        [84].runs[11] := 9, [84].runs[12] := 9, [84].runs[13] := 9, [84].runs[14] := 9, [84].runs[15] := 10, [84].runs[16] := 9, [84].runs[17] := 10, [84].runs[18] := 9, [84].runs[19] := 10, [84].runs[20] := 9, [84].runs[21] := 8, [84].runs[22] := 5, [84].time_avg[0] := 173, [84].time_avg[2] := 6434, [84].time_avg[3] := 9546, [84].time_avg[4] := 19840, [84].time_avg[5] := 19601, [84].time_avg[10] := 183, [84].time_avg[11] := 176, [84].time_avg[12] := 189, [84].time_avg[13] := 198, [84].time_avg[14] := 193, [84].time_avg[15] := 154, [84].time_avg[16] := 205, [84].time_avg[17] := 165, [84].time_avg[18] := 168, [84].time_avg[19] := 167, [84].time_avg[20] := 143, [84].time_avg[21] := 164, [84].time_avg[22] := 139, [85].date[0] := 19, [85].date[1] := 8, [85].date[2] := 23, [85].runs[0] := 108, [85].runs[7] := 1, [85].runs[9] := 4, [85].runs[10] := 3, [85].runs[11] := 10, [85].runs[12] := 9, [85].runs[13] := 8, [85].runs[14] := 9, [85].runs[15] := 10, [85].runs[16] := 9, [85].runs[17] := 9, [85].runs[18] := 8, [85].runs[19] := 9, [85].runs[20] := 9, [85].runs[21] := 8, [85].runs[22] := 2, [85].time_avg[0] := 204, [85].time_avg[2] := 6887, [85].time_avg[3] := 14477, [85].time_avg[4] := 20521, [85].time_avg[5] := 36240, [85].time_avg[10] := 221, [85].time_avg[11] := 190, [85].time_avg[12] := 186, [85].time_avg[13] := 191, [85].time_avg[14] := 226, [85].time_avg[15] := 161,
        [85].time_avg[16] := 185, [85].time_avg[17] := 211, [85].time_avg[18] := 232, [85].time_avg[19] := 218, [85].time_avg[20] := 196, [85].time_avg[21] := 251, [85].time_avg[22] := 235, [86].date[0] := 19, [86].date[1] := 8, [86].date[2] := 22, [86].runs[0] := 108, [86].runs[9] := 4, [86].runs[10] := 5, [86].runs[11] := 10, [86].runs[12] := 9, [86].runs[13] := 11, [86].runs[14] := 9, [86].runs[15] := 10, [86].runs[16] := 9, [86].runs[17] := 10, [86].runs[18] := 8, [86].runs[19] := 10, [86].runs[20] := 9, [86].runs[21] := 3, [86].time_avg[0] := 162, [86].time_avg[2] := 5022, [86].time_avg[3] := 11042, [86].time_avg[4] := 16840, [86].time_avg[5] := 22478, [86].time_avg[10] := 152, [86].time_avg[11] := 173, [86].time_avg[12] := 166, [86].time_avg[13] := 153, [86].time_avg[14] := 137, [86].time_avg[15] := 192, [86].time_avg[16] := 160, [86].time_avg[17] := 147, [86].time_avg[18] := 177, [86].time_avg[19] := 145, [86].time_avg[20] := 166, [86].time_avg[21] := 190, [87].date[0] := 19, [87].date[1] := 8, [87].date[2] := 21, [87].runs[0] := 110, [87].runs[9] := 5, [87].runs[10] := 5, [87].runs[11] := 9, [87].runs[12] := 8, [87].runs[13] := 10, [87].runs[14] := 10, [87].runs[15] := 10, [87].runs[16] := 10, [87].runs[17] := 9, [87].runs[18] := 10, [87].runs[19] := 8, [87].runs[20] := 9, [87].runs[21] := 6, [87].time_avg[0] := 174, [87].time_avg[2] := 5028,
        [87].time_avg[3] := 12622, [87].time_avg[4] := 18641, [87].time_avg[5] := 20757, [87].time_avg[9] := 267, [87].time_avg[10] := 158, [87].time_avg[11] := 186, [87].time_avg[12] := 162, [87].time_avg[13] := 179, [87].time_avg[14] := 156, [87].time_avg[15] := 147, [87].time_avg[16] := 154, [87].time_avg[17] := 158, [87].time_avg[18] := 185, [87].time_avg[19] := 180, [87].time_avg[20] := 236, [87].time_avg[21] := 167, [88].date[0] := 19, [88].date[1] := 8, [88].date[2] := 19, [88].runs[0] := 172, [88].runs[7] := 1, [88].runs[9] := 1, [88].runs[10] := 7, [88].runs[11] := 9, [88].runs[12] := 10, [88].runs[13] := 10, [88].runs[14] := 10, [88].runs[15] := 10, [88].runs[16] := 9, [88].runs[17] := 9, [88].runs[18] := 10, [88].runs[19] := 11, [88].runs[20] := 10, [88].runs[21] := 8, [88].time_avg[0] := 159, [88].time_avg[2] := 5010, [88].time_avg[3] := 9465, [88].time_avg[4] := 20080, [88].time_avg[5] := 17563, [88].time_avg[10] := 264, [88].time_avg[11] := 192, [88].time_avg[12] := 158, [88].time_avg[13] := 167, [88].time_avg[14] := 165, [88].time_avg[15] := 148, [88].time_avg[16] := 206, [88].time_avg[17] := 174, [88].time_avg[18] := 142, [88].time_avg[19] := 133, [88].time_avg[20] := 165, [88].time_avg[21] := 129, [89].date[0] := 19, [89].date[1] := 8, [89].date[2] := 18, [89].runs[0] := 116, [89].runs[7] := 1, [89].runs[10] := 8, [89].runs[11] := 10, [89].runs[12] := 10, [89].runs[13] := 9,
        [89].runs[14] := 10, [89].runs[15] := 11, [89].runs[16] := 4, [89].runs[17] := 9, [89].runs[18] := 10, [89].runs[19] := 10, [89].runs[20] := 9, [89].runs[21] := 11, [89].runs[22] := 4, [89].time_avg[0] := 160, [89].time_avg[2] := 4655, [89].time_avg[3] := 12877, [89].time_avg[4] := 21363, [89].time_avg[5] := 26439, [89].time_avg[10] := 166, [89].time_avg[11] := 166, [89].time_avg[12] := 161, [89].time_avg[13] := 187, [89].time_avg[14] := 165, [89].time_avg[15] := 133, [89].time_avg[16] := 160, [89].time_avg[17] := 161, [89].time_avg[18] := 173, [89].time_avg[19] := 149, [89].time_avg[20] := 175, [89].time_avg[21] := 139, [89].time_avg[22] := 162, [90].date[0] := 19, [90].date[1] := 8, [90].date[2] := 17, [90].runs[0] := 129, [90].runs[7] := 1, [90].runs[9] := 4, [90].runs[10] := 4, [90].runs[11] := 10, [90].runs[12] := 9, [90].runs[13] := 10, [90].runs[14] := 10, [90].runs[15] := 9, [90].runs[16] := 10, [90].runs[17] := 10, [90].runs[18] := 7, [90].runs[19] := 9, [90].runs[20] := 8, [90].runs[21] := 9, [90].runs[22] := 10, [90].runs[23] := 8, [90].time_avg[0] := 182, [90].time_avg[2] := 4196, [90].time_avg[3] := 11369, [90].time_avg[4] := 22122, [90].time_avg[5] := 21841, [90].time_avg[10] := 197, [90].time_avg[11] := 174, [90].time_avg[12] := 191, [90].time_avg[13] := 174, [90].time_avg[14] := 150, [90].time_avg[15] := 171, [90].time_avg[16] := 159, [90].time_avg[17] := 162,
        [90].time_avg[18] := 179, [90].time_avg[19] := 213, [90].time_avg[20] := 216, [90].time_avg[21] := 192, [90].time_avg[22] := 182, [90].time_avg[23] := 211, [91].date[0] := 19, [91].date[1] := 8, [91].date[2] := 16, [91].runs[0] := 110, [91].runs[7] := 1, [91].runs[9] := 4, [91].runs[10] := 6, [91].runs[11] := 10, [91].runs[12] := 8, [91].runs[13] := 9, [91].runs[14] := 3, [91].runs[15] := 10, [91].runs[16] := 10, [91].runs[17] := 10, [91].runs[18] := 9, [91].runs[19] := 9, [91].runs[20] := 9, [91].runs[21] := 10, [91].runs[22] := 2, [91].time_avg[0] := 167, [91].time_avg[2] := 5926, [91].time_avg[3] := 9632, [91].time_avg[4] := 23480, [91].time_avg[5] := 18838, [91].time_avg[10] := 161, [91].time_avg[11] := 149, [91].time_avg[12] := 156, [91].time_avg[13] := 170, [91].time_avg[15] := 151, [91].time_avg[16] := 156, [91].time_avg[17] := 158, [91].time_avg[18] := 203, [91].time_avg[19] := 192, [91].time_avg[20] := 185, [91].time_avg[21] := 150, [91].time_avg[22] := 195, [92].date[0] := 19, [92].date[1] := 8, [92].date[2] := 15, [92].runs[0] := 113, [92].runs[7] := 1, [92].runs[9] := 4, [92].runs[10] := 5, [92].runs[11] := 9, [92].runs[12] := 9, [92].runs[13] := 9, [92].runs[14] := 9, [92].runs[15] := 10, [92].runs[16] := 10, [92].runs[17] := 9, [92].runs[18] := 10, [92].runs[19] := 9, [92].runs[20] := 10, [92].runs[21] := 9,
        [92].time_avg[0] := 174, [92].time_avg[2] := 4980, [92].time_avg[3] := 11102, [92].time_avg[4] := 19122, [92].time_avg[5] := 22677, [92].time_avg[10] := 180, [92].time_avg[11] := 184, [92].time_avg[12] := 201, [92].time_avg[13] := 188, [92].time_avg[14] := 179, [92].time_avg[15] := 164, [92].time_avg[16] := 165, [92].time_avg[17] := 189, [92].time_avg[18] := 169, [92].time_avg[19] := 168, [92].time_avg[20] := 159, [92].time_avg[21] := 153, [93].date[0] := 19, [93].date[1] := 8, [93].date[2] := 14, [93].runs[0] := 110, [93].runs[7] := 1, [93].runs[9] := 4, [93].runs[10] := 5, [93].runs[11] := 9, [93].runs[12] := 10, [93].runs[13] := 10, [93].runs[14] := 10, [93].runs[15] := 10, [93].runs[16] := 10, [93].runs[17] := 8, [93].runs[18] := 10, [93].runs[19] := 10, [93].runs[20] := 8, [93].runs[21] := 5, [93].time_avg[0] := 170, [93].time_avg[2] := 3396, [93].time_avg[3] := 11574, [93].time_avg[4] := 19402, [93].time_avg[5] := 24403, [93].time_avg[10] := 164, [93].time_avg[11] := 183, [93].time_avg[12] := 161, [93].time_avg[13] := 163, [93].time_avg[14] := 151, [93].time_avg[15] := 150, [93].time_avg[16] := 168, [93].time_avg[17] := 227, [93].time_avg[18] := 179, [93].time_avg[19] := 161, [93].time_avg[20] := 173, [93].time_avg[21] := 178, [94].date[0] := 19, [94].date[1] := 8, [94].date[2] := 13, [94].runs[0] := 99, [94].runs[7] := 1, [94].runs[9] := 4, [94].runs[10] := 4, [94].runs[11] := 11,
        [94].runs[12] := 8, [94].runs[13] := 5, [94].runs[14] := 9, [94].runs[15] := 8, [94].runs[16] := 10, [94].runs[17] := 9, [94].runs[18] := 8, [94].runs[19] := 9, [94].runs[20] := 8, [94].runs[21] := 5, [94].time_avg[0] := 185, [94].time_avg[2] := 4905, [94].time_avg[3] := 9992, [94].time_avg[4] := 19077, [94].time_avg[5] := 20762, [94].time_avg[10] := 183, [94].time_avg[11] := 135, [94].time_avg[12] := 171, [94].time_avg[13] := 195, [94].time_avg[14] := 209, [94].time_avg[15] := 185, [94].time_avg[16] := 185, [94].time_avg[17] := 186, [94].time_avg[18] := 200, [94].time_avg[19] := 175, [94].time_avg[20] := 224, [94].time_avg[21] := 204, [95].date[0] := 19, [95].date[1] := 8, [95].date[2] := 12, [95].runs[0] := 118, [95].runs[8] := 1, [95].runs[9] := 6, [95].runs[10] := 5, [95].runs[11] := 10, [95].runs[12] := 11, [95].runs[13] := 10, [95].runs[14] := 8, [95].runs[15] := 10, [95].runs[16] := 10, [95].runs[17] := 10, [95].runs[18] := 10, [95].runs[19] := 8, [95].runs[20] := 9, [95].runs[21] := 10, [95].time_avg[0] := 156, [95].time_avg[2] := 6366, [95].time_avg[3] := 11660, [95].time_avg[4] := 23243, [95].time_avg[5] := 28239, [95].time_avg[10] := 194, [95].time_avg[11] := 153, [95].time_avg[12] := 133, [95].time_avg[13] := 156, [95].time_avg[14] := 137, [95].time_avg[15] := 150, [95].time_avg[16] := 151, [95].time_avg[17] := 145, [95].time_avg[18] := 164, [95].time_avg[19] := 182,
        [95].time_avg[20] := 195, [95].time_avg[21] := 148, [96].date[0] := 19, [96].date[1] := 8, [96].date[2] := 11, [96].runs[0] := 123, [96].runs[7] := 1, [96].runs[9] := 4, [96].runs[10] := 8, [96].runs[11] := 10, [96].runs[12] := 11, [96].runs[13] := 10, [96].runs[14] := 7, [96].runs[15] := 11, [96].runs[16] := 9, [96].runs[17] := 10, [96].runs[18] := 9, [96].runs[19] := 11, [96].runs[20] := 8, [96].runs[21] := 9, [96].runs[22] := 5, [96].time_avg[0] := 157, [96].time_avg[2] := 4752, [96].time_avg[3] := 9692, [96].time_avg[4] := 19361, [96].time_avg[5] := 22281, [96].time_avg[10] := 173, [96].time_avg[11] := 141, [96].time_avg[12] := 142, [96].time_avg[13] := 141, [96].time_avg[14] := 179, [96].time_avg[15] := 138, [96].time_avg[16] := 183, [96].time_avg[17] := 147, [96].time_avg[18] := 191, [96].time_avg[19] := 146, [96].time_avg[20] := 167, [96].time_avg[21] := 162, [96].time_avg[22] := 167, [97].date[0] := 19, [97].date[1] := 8, [97].date[2] := 10, [97].runs[0] := 120, [97].runs[7] := 1, [97].runs[9] := 5, [97].runs[10] := 4, [97].runs[11] := 6, [97].runs[12] := 8, [97].runs[13] := 11, [97].runs[14] := 8, [97].runs[15] := 11, [97].runs[16] := 9, [97].runs[17] := 10, [97].runs[18] := 11, [97].runs[19] := 10, [97].runs[20] := 11, [97].runs[21] := 10, [97].runs[22] := 5, [97].time_avg[0] := 142, [97].time_avg[2] := 4697,
        [97].time_avg[3] := 8479, [97].time_avg[4] := 21362, [97].time_avg[5] := 36560, [97].time_avg[10] := 200, [97].time_avg[11] := 178, [97].time_avg[12] := 152, [97].time_avg[13] := 141, [97].time_avg[14] := 131, [97].time_avg[15] := 153, [97].time_avg[16] := 133, [97].time_avg[17] := 145, [97].time_avg[18] := 140, [97].time_avg[19] := 135, [97].time_avg[20] := 138, [97].time_avg[21] := 126, [97].time_avg[22] := 121, [98].date[0] := 19, [98].date[1] := 8, [98].date[2] := 9, [98].runs[0] := 119, [98].runs[7] := 1, [98].runs[9] := 5, [98].runs[10] := 5, [98].runs[11] := 8, [98].runs[12] := 9, [98].runs[13] := 8, [98].runs[14] := 11, [98].runs[15] := 11, [98].runs[16] := 8, [98].runs[17] := 10, [98].runs[18] := 9, [98].runs[19] := 11, [98].runs[20] := 9, [98].runs[21] := 10, [98].runs[22] := 4, [98].time_avg[0] := 151, [98].time_avg[2] := 4804, [98].time_avg[3] := 10881, [98].time_avg[4] := 800, [98].time_avg[5] := 21920, [98].time_avg[9] := 35, [98].time_avg[10] := 126, [98].time_avg[11] := 166, [98].time_avg[12] := 159, [98].time_avg[13] := 165, [98].time_avg[14] := 138, [98].time_avg[15] := 126, [98].time_avg[16] := 148, [98].time_avg[17] := 148, [98].time_avg[18] := 187, [98].time_avg[19] := 138, [98].time_avg[20] := 165, [98].time_avg[21] := 145, [98].time_avg[22] := 168, [99].date[0] := 19, [99].date[1] := 8, [99].date[2] := 8, [99].runs[0] := 93, [99].runs[7] := 1, [99].runs[9] := 4,
        [99].runs[10] := 4, [99].runs[11] := 9, [99].runs[12] := 9, [99].runs[13] := 9, [99].runs[14] := 8, [99].runs[15] := 9, [99].runs[16] := 9, [99].runs[17] := 2, [99].runs[18] := 5, [99].runs[19] := 8, [99].runs[20] := 9, [99].runs[21] := 7, [99].time_avg[0] := 156, [99].time_avg[2] := 5998, [99].time_avg[3] := 7111, [99].time_avg[4] := 17880, [99].time_avg[5] := 21321, [99].time_avg[10] := 153, [99].time_avg[11] := 154, [99].time_avg[12] := 146, [99].time_avg[13] := 139, [99].time_avg[14] := 173, [99].time_avg[15] := 152, [99].time_avg[16] := 160, [99].time_avg[17] := 133, [99].time_avg[18] := 182, [99].time_avg[19] := 147, [99].time_avg[20] := 148, [99].time_avg[21] := 188);
        [0].time_avg[2]   // Daily Avg Platform Cycle Waiting After Cycle
        [0].time_avg[3]   // Daily Avg Platform Cycle Before Start Cycle
        [0].time_avg[4]   // Overall Time End of Cycle Plat
        [0].time_avg[5]   // Overall Time Before Cycle Plat
   JM_Statistics_Storage : Run_Count_Hist_JM[100] := ([1].date[0] := 25, [1].date[1] := 11, [1].date[2] := 28, [1].runs[0] := 65, [1].runs[8] := 2, [1].runs[9] := 1, [1].runs[15] := 3, [1].runs[16] := 7, [1].runs[17] := 8, [1].runs[18] := 8, [1].runs[19] := 8, [1].runs[20] := 8, [1].runs[21] := 7, [1].runs[22] := 8, [1].runs[23] := 5, [1].time_avg[0] := 204, [1].time_avg[2] := 3400, [1].time_avg[4] := 19639, [1].time_avg[5] := 22361, [1].time_avg[8] := 50, [1].time_avg[15] := 203, [1].time_avg[16] := 254, [1].time_avg[17] := 210, [1].time_avg[18] := 202, [1].time_avg[19] := 195, [1].time_avg[20] := 206, [1].time_avg[21] := 190, [1].time_avg[22] := 211, [1].time_avg[23] := 177, [2].date[0] := 25, [2].date[1] := 11, [2].date[2] := 27, [2].runs[0] := 63, [2].runs[14] := 6, [2].runs[15] := 4, [2].runs[16] := 7, [2].runs[17] := 7, [2].runs[18] := 8, [2].runs[19] := 8, [2].runs[20] := 7, [2].runs[21] := 5, [2].runs[22] := 8, [2].runs[23] := 3, [2].time_avg[0] := 234, [2].time_avg[4] := 21760, [2].time_avg[5] := 22361, [2].time_avg[14] := 167, [2].time_avg[15] := 316, [2].time_avg[16] := 272, [2].time_avg[17] := 206, [2].time_avg[18] := 208, [2].time_avg[19] := 242, [2].time_avg[20] := 266, [2].time_avg[21] := 233, [2].time_avg[22] := 223, [2].time_avg[23] := 245, [3].date[0] := 25, [3].date[1] := 11, [3].date[2] := 26, [3].runs[0] := 57,
        [3].runs[12] := 4, [3].runs[13] := 1, [3].runs[15] := 2, [3].runs[16] := 6, [3].runs[17] := 7, [3].runs[18] := 7, [3].runs[19] := 7, [3].runs[20] := 7, [3].runs[21] := 7, [3].runs[22] := 6, [3].runs[23] := 3, [3].time_avg[0] := 274, [3].time_avg[2] := 6041, [3].time_avg[4] := 21760, [3].time_avg[5] := 22361, [3].time_avg[12] := 396, [3].time_avg[13] := 320, [3].time_avg[15] := 271, [3].time_avg[16] := 271, [3].time_avg[17] := 292, [3].time_avg[18] := 243, [3].time_avg[19] := 255, [3].time_avg[20] := 243, [3].time_avg[21] := 289, [3].time_avg[22] := 278, [3].time_avg[23] := 283, [4].date[0] := 25, [4].date[1] := 11, [4].date[2] := 25, [4].runs[0] := 53, [4].runs[7] := 1, [4].runs[15] := 1, [4].runs[16] := 5, [4].runs[17] := 8, [4].runs[18] := 6, [4].runs[19] := 8, [4].runs[20] := 7, [4].runs[21] := 7, [4].runs[22] := 7, [4].runs[23] := 3, [4].time_avg[0] := 260, [4].time_avg[4] := 53080, [4].time_avg[5] := 22361, [4].time_avg[16] := 223, [4].time_avg[17] := 286, [4].time_avg[18] := 280, [4].time_avg[19] := 258, [4].time_avg[20] := 261, [4].time_avg[21] := 234, [4].time_avg[22] := 267, [4].time_avg[23] := 254, [5].date[0] := 25, [5].date[1] := 11, [5].date[2] := 24, [5].runs[0] := 67, [5].runs[7] := 4, [5].runs[8] := 3, [5].runs[10] := 2, [5].runs[11] := 4, [5].runs[13] := 1,
        [5].runs[14] := 1, [5].runs[15] := 4, [5].runs[16] := 7, [5].runs[17] := 7, [5].runs[18] := 7, [5].runs[19] := 7, [5].runs[20] := 4, [5].runs[21] := 7, [5].runs[22] := 6, [5].runs[23] := 3, [5].time_avg[0] := 254, [5].time_avg[2] := 76642, [5].time_avg[4] := 53080, [5].time_avg[5] := 22361, [5].time_avg[7] := 75, [5].time_avg[8] := 246, [5].time_avg[11] := 171, [5].time_avg[14] := 83, [5].time_avg[15] := 147, [5].time_avg[16] := 272, [5].time_avg[17] := 276, [5].time_avg[18] := 244, [5].time_avg[19] := 256, [5].time_avg[20] := 266, [5].time_avg[21] := 291, [5].time_avg[22] := 291, [5].time_avg[23] := 290, [6].date[0] := 25, [6].date[1] := 11, [6].date[2] := 23, [6].runs[0] := 54, [6].runs[10] := 2, [6].runs[11] := 4, [6].runs[15] := 1, [6].runs[16] := 8, [6].runs[17] := 7, [6].runs[18] := 6, [6].runs[19] := 5, [6].runs[20] := 8, [6].runs[21] := 6, [6].runs[22] := 5, [6].runs[23] := 2, [6].time_avg[0] := 268, [6].time_avg[4] := 23760, [6].time_avg[5] := 22361, [6].time_avg[11] := 332, [6].time_avg[16] := 211, [6].time_avg[17] := 253, [6].time_avg[18] := 262, [6].time_avg[19] := 274, [6].time_avg[20] := 241, [6].time_avg[21] := 295, [6].time_avg[22] := 310, [6].time_avg[23] := 371, [7].date[0] := 25, [7].date[1] := 11, [7].date[2] := 22, [7].runs[0] := 49, [7].runs[12] := 7, [7].runs[14] := 1,
        [7].runs[15] := 4, [7].runs[16] := 7, [7].runs[17] := 7, [7].runs[18] := 7, [7].runs[19] := 1, [7].runs[20] := 6, [7].runs[21] := 2, [7].runs[22] := 6, [7].runs[23] := 1, [7].time_avg[0] := 278, [7].time_avg[4] := 23760, [7].time_avg[5] := 22361, [7].time_avg[12] := 180, [7].time_avg[15] := 308, [7].time_avg[16] := 282, [7].time_avg[17] := 261, [7].time_avg[18] := 280, [7].time_avg[19] := 295, [7].time_avg[20] := 361, [7].time_avg[22] := 287, [8].date[0] := 25, [8].date[1] := 11, [8].date[2] := 20, [8].runs[0] := 58, [8].runs[10] := 2, [8].runs[11] := 3, [8].runs[13] := 5, [8].runs[14] := 4, [8].runs[15] := 3, [8].runs[16] := 5, [8].runs[17] := 4, [8].runs[18] := 3, [8].runs[19] := 6, [8].runs[20] := 5, [8].runs[21] := 7, [8].runs[22] := 7, [8].runs[23] := 4, [8].time_avg[0] := 205, [8].time_avg[2] := 15381, [8].time_avg[4] := 23760, [8].time_avg[5] := 22361, [8].time_avg[10] := 76, [8].time_avg[11] := 152, [8].time_avg[13] := 198, [8].time_avg[14] := 60, [8].time_avg[15] := 73, [8].time_avg[16] := 76, [8].time_avg[17] := 183, [8].time_avg[18] := 376, [8].time_avg[19] := 286, [8].time_avg[20] := 250, [8].time_avg[21] := 218, [8].time_avg[22] := 239, [8].time_avg[23] := 211, [9].date[0] := 25, [9].date[1] := 11, [9].date[2] := 19, [9].runs[0] := 7, [9].runs[12] := 2, [9].runs[13] := 4,
        [9].runs[17] := 1, [9].runs[18] := 1, [9].time_avg[0] := 217, [9].time_avg[2] := 78801, [9].time_avg[4] := 48480, [9].time_avg[5] := 22361, [9].time_avg[13] := 217, [10].date[0] := 25, [10].date[1] := 11, [10].date[2] := 16, [10].runs[0] := 7, [10].runs[10] := 2, [10].runs[13] := 7, [10].time_avg[0] := 93, [10].time_avg[4] := 27759, [10].time_avg[5] := 22361, [10].time_avg[13] := 93, [11].date[0] := 25, [11].date[1] := 11, [11].date[2] := 14, [11].runs[0] := 2, [11].runs[15] := 1, [11].runs[16] := 1, [11].time_avg[2] := 32760, [11].time_avg[4] := 27759, [11].time_avg[5] := 22361, [12].date[0] := 25, [12].date[1] := 11, [12].date[2] := 13, [12].runs[0] := 14, [12].runs[10] := 2, [12].runs[11] := 1, [12].runs[12] := 1, [12].runs[14] := 2, [12].runs[15] := 5, [12].runs[16] := 4, [12].runs[17] := 5, [12].time_avg[0] := 141, [12].time_avg[4] := 36240, [12].time_avg[5] := 22361, [12].time_avg[10] := 210, [12].time_avg[14] := 205, [12].time_avg[15] := 160, [12].time_avg[16] := 100, [12].time_avg[17] := 100, [13].date[0] := 25, [13].date[1] := 11, [13].date[2] := 11, [13].runs[0] := 2, [13].runs[18] := 2, [13].time_avg[0] := 88, [13].time_avg[4] := 36240, [13].time_avg[5] := 22361, [13].time_avg[18] := 88, [14].date[0] := 25, [14].date[1] := 11, [14].date[2] := 7, [14].runs[0] := 5, [14].runs[15] := 3, [14].runs[16] := 2,
        [14].time_avg[0] := 229, [14].time_avg[4] := 36240, [14].time_avg[5] := 22361, [14].time_avg[15] := 300, [14].time_avg[16] := 87, [15].date[0] := 25, [15].date[1] := 11, [15].date[2] := 6, [15].runs[0] := 13, [15].runs[15] := 1, [15].runs[16] := 3, [15].runs[17] := 8, [15].runs[18] := 1, [15].runs[19] := 4, [15].time_avg[0] := 54, [15].time_avg[4] := 36240, [15].time_avg[5] := 22361, [15].time_avg[17] := 46, [15].time_avg[19] := 66, [16].date[0] := 25, [16].date[1] := 10, [16].date[2] := 27, [16].runs[0] := 13, [16].runs[12] := 1, [16].runs[13] := 4, [16].runs[14] := 1, [16].time_avg[0] := 126, [16].time_avg[4] := 36240, [16].time_avg[5] := 22361, [16].time_avg[13] := 65, [17].date[0] := 25, [17].date[1] := 10, [17].date[2] := 26, [17].runs[0] := 58, [17].runs[10] := 1, [17].runs[11] := 2, [17].runs[12] := 3, [17].runs[13] := 8, [17].runs[14] := 8, [17].runs[15] := 6, [17].runs[16] := 7, [17].runs[17] := 7, [17].runs[18] := 6, [17].runs[19] := 7, [17].runs[20] := 3, [17].time_avg[0] := 252, [17].time_avg[2] := 40720, [17].time_avg[4] := 36240, [17].time_avg[5] := 22361, [17].time_avg[11] := 476, [17].time_avg[12] := 190, [17].time_avg[13] := 206, [17].time_avg[14] := 216, [17].time_avg[15] := 310, [17].time_avg[16] := 261, [17].time_avg[17] := 248, [17].time_avg[18] := 232, [17].time_avg[19] := 304, [17].time_avg[20] := 214, [18].date[0] := 25,
        [18].date[1] := 10, [18].date[2] := 25, [18].runs[0] := 47, [18].runs[12] := 5, [18].runs[13] := 9, [18].runs[14] := 5, [18].runs[16] := 2, [18].runs[17] := 8, [18].runs[18] := 7, [18].runs[19] := 7, [18].runs[20] := 4, [18].time_avg[0] := 227, [18].time_avg[4] := 26040, [18].time_avg[5] := 22361, [18].time_avg[12] := 203, [18].time_avg[13] := 166, [18].time_avg[14] := 231, [18].time_avg[16] := 370, [18].time_avg[17] := 239, [18].time_avg[18] := 252, [18].time_avg[19] := 244, [18].time_avg[20] := 235, [19].date[0] := 25, [19].date[1] := 10, [19].date[2] := 23, [19].runs[0] := 48, [19].runs[9] := 2, [19].runs[10] := 3, [19].runs[12] := 3, [19].runs[13] := 7, [19].runs[14] := 7, [19].runs[15] := 5, [19].runs[16] := 8, [19].runs[17] := 5, [19].runs[19] := 5, [19].runs[20] := 3, [19].time_avg[0] := 257, [19].time_avg[2] := 18201, [19].time_avg[4] := 26040, [19].time_avg[5] := 22361, [19].time_avg[9] := 102, [19].time_avg[10] := 259, [19].time_avg[12] := 493, [19].time_avg[13] := 241, [19].time_avg[14] := 231, [19].time_avg[15] := 264, [19].time_avg[16] := 252, [19].time_avg[17] := 280, [19].time_avg[19] := 300, [19].time_avg[20] := 235, [20].date[0] := 25, [20].date[1] := 10, [20].date[2] := 22, [20].runs[0] := 62, [20].runs[10] := 4, [20].runs[12] := 2, [20].runs[13] := 9, [20].runs[14] := 7, [20].runs[15] := 7, [20].runs[16] := 7,
        [20].runs[17] := 7, [20].runs[18] := 8, [20].runs[19] := 8, [20].runs[20] := 3, [20].time_avg[0] := 226, [20].time_avg[4] := 26079, [20].time_avg[5] := 22361, [20].time_avg[10] := 123, [20].time_avg[13] := 199, [20].time_avg[14] := 230, [20].time_avg[15] := 230, [20].time_avg[16] := 312, [20].time_avg[17] := 253, [20].time_avg[18] := 219, [20].time_avg[19] := 200, [20].time_avg[20] := 206, [21].date[0] := 25, [21].date[1] := 10, [21].date[2] := 21, [21].runs[0] := 58, [21].runs[11] := 3, [21].runs[12] := 1, [21].runs[13] := 8, [21].runs[14] := 7, [21].runs[15] := 4, [21].runs[16] := 8, [21].runs[17] := 8, [21].runs[18] := 7, [21].runs[19] := 8, [21].runs[20] := 4, [21].time_avg[0] := 233, [21].time_avg[2] := 42160, [21].time_avg[4] := 26079, [21].time_avg[5] := 22361, [21].time_avg[11] := 186, [21].time_avg[13] := 222, [21].time_avg[14] := 240, [21].time_avg[15] := 294, [21].time_avg[16] := 256, [21].time_avg[17] := 202, [21].time_avg[18] := 246, [21].time_avg[19] := 216, [21].time_avg[20] := 208, [22].date[0] := 25, [22].date[1] := 10, [22].date[2] := 20, [22].runs[0] := 47, [22].runs[10] := 2, [22].runs[11] := 6, [22].runs[12] := 1, [22].runs[13] := 7, [22].runs[14] := 7, [22].runs[15] := 7, [22].runs[16] := 4, [22].runs[17] := 1, [22].runs[18] := 2, [22].runs[19] := 7, [22].runs[20] := 3, [22].time_avg[0] := 249, [22].time_avg[2] := 52640,
        [22].time_avg[4] := 40960, [22].time_avg[5] := 22361, [22].time_avg[11] := 232, [22].time_avg[13] := 215, [22].time_avg[14] := 258, [22].time_avg[15] := 237, [22].time_avg[16] := 210, [22].time_avg[18] := 331, [22].time_avg[19] := 294, [22].time_avg[20] := 241, [23].date[0] := 25, [23].date[1] := 10, [23].date[2] := 19, [23].runs[0] := 61, [23].runs[9] := 2, [23].runs[10] := 2, [23].runs[11] := 8, [23].runs[12] := 4, [23].runs[13] := 6, [23].runs[14] := 1, [23].runs[15] := 8, [23].runs[16] := 7, [23].runs[17] := 7, [23].runs[18] := 7, [23].runs[19] := 7, [23].runs[20] := 2, [23].time_avg[0] := 237, [23].time_avg[2] := 59762, [23].time_avg[4] := 52320, [23].time_avg[5] := 22361, [23].time_avg[9] := 89, [23].time_avg[11] := 203, [23].time_avg[12] := 193, [23].time_avg[13] := 194, [23].time_avg[15] := 243, [23].time_avg[16] := 238, [23].time_avg[17] := 251, [23].time_avg[18] := 268, [23].time_avg[19] := 280, [23].time_avg[20] := 287, [24].date[0] := 25, [24].date[1] := 10, [24].date[2] := 18, [24].runs[0] := 51, [24].runs[9] := 2, [24].runs[10] := 5, [24].runs[11] := 8, [24].runs[12] := 2, [24].runs[13] := 5, [24].runs[14] := 6, [24].runs[15] := 7, [24].runs[16] := 5, [24].runs[17] := 7, [24].runs[18] := 4, [24].time_avg[0] := 246, [24].time_avg[4] := 52360, [24].time_avg[5] := 22361, [24].time_avg[10] := 182, [24].time_avg[11] := 228, [24].time_avg[12] := 212,
        [24].time_avg[13] := 231, [24].time_avg[14] := 324, [24].time_avg[15] := 255, [24].time_avg[16] := 238, [24].time_avg[17] := 263, [24].time_avg[18] := 255, [25].date[0] := 25, [25].date[1] := 10, [25].date[2] := 15, [25].runs[0] := 89, [25].runs[10] := 4, [25].runs[11] := 4, [25].runs[12] := 7, [25].runs[13] := 6, [25].runs[14] := 8, [25].runs[15] := 6, [25].runs[16] := 7, [25].runs[17] := 6, [25].time_avg[0] := 251, [25].time_avg[2] := 50482, [25].time_avg[4] := 52360, [25].time_avg[5] := 22361, [25].time_avg[10] := 61, [25].time_avg[11] := 214, [25].time_avg[12] := 261, [25].time_avg[13] := 348, [25].time_avg[14] := 197, [25].time_avg[15] := 264, [25].time_avg[16] := 241, [25].time_avg[17] := 309, [26].date[0] := 25, [26].date[1] := 10, [26].date[2] := 14, [26].runs[0] := 14, [26].runs[10] := 5, [26].runs[11] := 1, [26].runs[12] := 8, [26].time_avg[0] := 175, [26].time_avg[4] := 34119, [26].time_avg[5] := 22361, [26].time_avg[10] := 270, [26].time_avg[12] := 121, [27].date[0] := 25, [27].date[1] := 10, [27].date[2] := 13, [27].runs[0] := 29, [27].runs[12] := 3, [27].runs[13] := 5, [27].runs[14] := 6, [27].runs[15] := 4, [27].runs[16] := 7, [27].runs[17] := 4, [27].time_avg[0] := 256, [27].time_avg[2] := 63880, [27].time_avg[4] := 34119, [27].time_avg[5] := 22361, [27].time_avg[12] := 68, [27].time_avg[13] := 218, [27].time_avg[14] := 246, [27].time_avg[15] := 367,
        [27].time_avg[16] := 315, [27].time_avg[17] := 255, [28].date[0] := 25, [28].date[1] := 10, [28].date[2] := 10, [28].runs[0] := 27, [28].runs[9] := 9, [28].runs[10] := 11, [28].runs[11] := 7, [28].time_avg[0] := 89, [28].time_avg[4] := 33481, [28].time_avg[5] := 22361, [28].time_avg[9] := 82, [28].time_avg[10] := 83, [28].time_avg[11] := 123, [29].date[0] := 25, [29].date[1] := 10, [29].date[2] := 8, [29].runs[0] := 76, [29].runs[9] := 9, [29].runs[10] := 11, [29].runs[11] := 8, [29].runs[12] := 10, [29].runs[13] := 11, [29].runs[14] := 7, [29].runs[15] := 7, [29].runs[16] := 3, [29].time_avg[0] := 100, [29].time_avg[4] := 33481, [29].time_avg[5] := 22361, [29].time_avg[9] := 47, [29].time_avg[10] := 77, [29].time_avg[11] := 96, [29].time_avg[12] := 96, [29].time_avg[13] := 82, [29].time_avg[14] := 70, [29].time_avg[15] := 221, [29].time_avg[16] := 56, [30].date[0] := 25, [30].date[1] := 10, [30].date[2] := 7, [30].runs[0] := 1, [30].runs[8] := 1, [30].time_avg[4] := 33481, [30].time_avg[5] := 22361, [31].date[0] := 25, [31].date[1] := 10, [31].date[2] := 6, [31].runs[0] := 3, [31].runs[12] := 3, [31].time_avg[0] := 51, [31].time_avg[4] := 33481, [31].time_avg[5] := 22361, [31].time_avg[12] := 51, [32].date[0] := 25, [32].date[1] := 10, [32].date[2] := 5, [32].runs[0] := 3, [32].runs[12] := 1, [32].runs[15] := 2,
        [32].time_avg[0] := 43, [32].time_avg[4] := 33481, [32].time_avg[5] := 22361, [32].time_avg[15] := 43, [33].date[0] := 25, [33].date[1] := 10, [33].date[2] := 4, [33].runs[0] := 15, [33].runs[10] := 4, [33].runs[11] := 3, [33].runs[12] := 3, [33].runs[15] := 4, [33].runs[16] := 1, [33].time_avg[0] := 228, [33].time_avg[2] := 47342, [33].time_avg[4] := 33481, [33].time_avg[5] := 22361, [33].time_avg[10] := 258, [33].time_avg[11] := 342, [33].time_avg[12] := 69, [33].time_avg[15] := 112, [34].date[0] := 25, [34].date[1] := 10, [34].date[2] := 1, [34].runs[0] := 64, [34].runs[9] := 1, [34].runs[10] := 7, [34].runs[11] := 8, [34].runs[12] := 9, [34].runs[13] := 6, [34].runs[14] := 8, [34].runs[15] := 9, [34].runs[16] := 8, [34].runs[17] := 8, [34].time_avg[0] := 168, [34].time_avg[4] := 53200, [34].time_avg[5] := 22361, [34].time_avg[10] := 151, [34].time_avg[11] := 172, [34].time_avg[12] := 168, [34].time_avg[13] := 171, [34].time_avg[14] := 150, [34].time_avg[15] := 177, [34].time_avg[16] := 175, [34].time_avg[17] := 175, [35].date[0] := 25, [35].date[1] := 9, [35].date[2] := 30, [35].runs[0] := 60, [35].runs[9] := 5, [35].runs[10] := 5, [35].runs[11] := 9, [35].runs[12] := 7, [35].runs[13] := 8, [35].runs[14] := 9, [35].runs[15] := 9, [35].runs[16] := 8, [35].time_avg[0] := 176, [35].time_avg[2] := 40561, [35].time_avg[4] := 53200,
        [35].time_avg[5] := 22361, [35].time_avg[9] := 120, [35].time_avg[10] := 150, [35].time_avg[11] := 176, [35].time_avg[12] := 186, [35].time_avg[13] := 219, [35].time_avg[14] := 153, [35].time_avg[15] := 180, [35].time_avg[16] := 165, [36].date[0] := 25, [36].date[1] := 9, [36].date[2] := 29, [36].runs[0] := 57, [36].runs[8] := 2, [36].runs[9] := 7, [36].runs[10] := 7, [36].runs[11] := 8, [36].runs[12] := 5, [36].runs[13] := 7, [36].runs[14] := 7, [36].runs[15] := 7, [36].runs[16] := 7, [36].time_avg[0] := 211, [36].time_avg[4] := 56839, [36].time_avg[5] := 22361, [36].time_avg[9] := 166, [36].time_avg[10] := 267, [36].time_avg[11] := 147, [36].time_avg[12] := 241, [36].time_avg[13] := 205, [36].time_avg[14] := 168, [36].time_avg[15] := 266, [36].time_avg[16] := 222, [37].date[0] := 25, [37].date[1] := 9, [37].date[2] := 28, [37].runs[0] := 58, [37].runs[9] := 3, [37].runs[10] := 9, [37].runs[11] := 7, [37].runs[12] := 8, [37].runs[13] := 8, [37].runs[14] := 8, [37].runs[15] := 7, [37].runs[16] := 8, [37].time_avg[0] := 184, [37].time_avg[4] := 56839, [37].time_avg[5] := 22361, [37].time_avg[9] := 167, [37].time_avg[10] := 193, [37].time_avg[11] := 208, [37].time_avg[12] := 169, [37].time_avg[13] := 199, [37].time_avg[14] := 199, [37].time_avg[15] := 173, [37].time_avg[16] := 151, [38].date[0] := 25, [38].date[1] := 9, [38].date[2] := 25, [38].runs[0] := 64,
        [38].runs[8] := 4, [38].runs[9] := 6, [38].runs[10] := 7, [38].runs[11] := 7, [38].runs[12] := 8, [38].runs[13] := 8, [38].runs[14] := 8, [38].runs[15] := 9, [38].runs[16] := 7, [38].time_avg[0] := 201, [38].time_avg[4] := 56839, [38].time_avg[5] := 22361, [38].time_avg[8] := 455, [38].time_avg[9] := 193, [38].time_avg[10] := 212, [38].time_avg[11] := 189, [38].time_avg[12] := 207, [38].time_avg[13] := 224, [38].time_avg[14] := 191, [38].time_avg[15] := 166, [38].time_avg[16] := 193, [39].date[0] := 25, [39].date[1] := 9, [39].date[2] := 24, [39].runs[0] := 50, [39].runs[9] := 4, [39].runs[10] := 6, [39].runs[11] := 5, [39].runs[12] := 6, [39].runs[13] := 5, [39].runs[14] := 8, [39].runs[15] := 8, [39].runs[16] := 8, [39].time_avg[0] := 195, [39].time_avg[4] := 56839, [39].time_avg[5] := 22361, [39].time_avg[9] := 83, [39].time_avg[10] := 198, [39].time_avg[11] := 260, [39].time_avg[12] := 133, [39].time_avg[13] := 207, [39].time_avg[14] := 244, [39].time_avg[15] := 215, [39].time_avg[16] := 169, [40].date[0] := 25, [40].date[1] := 9, [40].date[2] := 22, [40].runs[0] := 46, [40].runs[8] := 4, [40].runs[9] := 3, [40].runs[10] := 7, [40].runs[11] := 5, [40].runs[12] := 7, [40].runs[13] := 5, [40].runs[14] := 2, [40].runs[15] := 6, [40].runs[16] := 7, [40].time_avg[0] := 229, [40].time_avg[4] := 56839, [40].time_avg[5] := 22361,
        [40].time_avg[8] := 208, [40].time_avg[10] := 179, [40].time_avg[11] := 196, [40].time_avg[12] := 160, [40].time_avg[13] := 227, [40].time_avg[15] := 325, [40].time_avg[16] := 281, [41].date[0] := 25, [41].date[1] := 9, [41].date[2] := 21, [41].runs[0] := 9, [41].runs[8] := 1, [41].runs[9] := 6, [41].runs[14] := 2, [41].time_avg[0] := 233, [41].time_avg[2] := 43360, [41].time_avg[4] := 56839, [41].time_avg[5] := 22361, [41].time_avg[9] := 244, [41].time_avg[14] := 175, [42].date[0] := 25, [42].date[1] := 9, [42].date[2] := 18, [42].runs[0] := 6, [42].runs[11] := 5, [42].runs[12] := 1, [42].time_avg[0] := 226, [42].time_avg[4] := 37320, [42].time_avg[5] := 22361, [42].time_avg[11] := 226, [43].date[0] := 25, [43].date[1] := 9, [43].date[2] := 16, [43].runs[0] := 2, [43].runs[15] := 1, [43].runs[16] := 1, [43].time_avg[2] := 46801, [43].time_avg[4] := 37320, [43].time_avg[5] := 22361, [44].date[0] := 25, [44].date[1] := 8, [44].date[2] := 15, [44].runs[0] := 3, [44].runs[12] := 1, [44].runs[15] := 2, [44].time_avg[4] := 37641, [44].time_avg[5] := 22361, [45].date[0] := 25, [45].date[1] := 7, [45].date[2] := 13, [45].runs[0] := 107, [45].runs[9] := 2, [45].runs[14] := 2, [45].runs[16] := 8, [45].time_avg[0] := 162, [45].time_avg[2] := 22208, [45].time_avg[4] := 37641, [45].time_avg[5] := 22361, [45].time_avg[9] := 55, [45].time_avg[14] := 220,
        [45].time_avg[16] := 142, [46].date[0] := -2, [46].date[1] := 1, [46].date[2] := 15, [46].runs[0] := 1, [46].time_avg[4] := 45599, [46].time_avg[5] := 22361, [47].date[0] := -2, [47].date[1] := 1, [47].date[2] := 12, [47].runs[0] := 14, [47].runs[23] := 3, [47].time_avg[0] := 172, [47].time_avg[4] := 45599, [47].time_avg[5] := 22361, [47].time_avg[23] := 108, [48].date[0] := -2, [48].date[1] := 1, [48].date[2] := 11, [48].runs[0] := 14, [48].runs[21] := 1, [48].time_avg[0] := 145, [48].time_avg[4] := 45599, [48].time_avg[5] := 22361, [49].date[0] := -2, [49].date[1] := 1, [49].date[2] := 10, [49].runs[0] := 2, [49].runs[20] := 1, [49].runs[23] := 1, [49].time_avg[4] := 45599, [49].time_avg[5] := 22361, [50].date[0] := -2, [50].date[1] := 1, [50].date[2] := 8, [50].runs[0] := 1, [50].time_avg[4] := 45599, [50].time_avg[5] := 22361, [51].date[0] := -2, [51].date[1] := 1, [51].date[2] := 6, [51].runs[0] := 2, [51].runs[20] := 1, [51].time_avg[4] := 45599, [51].time_avg[5] := 22361, [52].date[0] := -2, [52].date[1] := 1, [52].date[2] := 5, [52].runs[0] := 10, [52].runs[20] := 2, [52].runs[23] := 3, [52].time_avg[0] := 139, [52].time_avg[4] := 45599, [52].time_avg[5] := 22361, [52].time_avg[23] := 139, [53].date[0] := -2, [53].date[1] := 1, [53].date[2] := 4, [53].runs[0] := 7, [53].runs[21] := 1,
        [53].runs[22] := 2, [53].time_avg[0] := 542, [53].time_avg[4] := 45599, [53].time_avg[5] := 22361, [53].time_avg[22] := 542, [54].date[0] := -2, [54].date[1] := 1, [54].date[2] := 2, [54].runs[0] := 4, [54].runs[23] := 4, [54].time_avg[4] := 45599, [54].time_avg[5] := 22361, [55].date[0] := -2, [55].date[1] := 1, [55].date[2] := 21, [55].runs[0] := 12, [55].runs[19] := 1, [55].runs[20] := 1, [55].runs[23] := 2, [55].time_avg[0] := 325, [55].time_avg[4] := 45599, [55].time_avg[5] := 22361, [56].date[0] := -2, [56].date[1] := 1, [56].date[2] := 20, [56].runs[0] := 15, [56].runs[17] := 4, [56].runs[18] := 1, [56].runs[23] := 1, [56].time_avg[0] := 214, [56].time_avg[2] := 35440, [56].time_avg[4] := 45599, [56].time_avg[5] := 22361, [56].time_avg[17] := 368, [57].date[0] := -2, [57].date[1] := 1, [57].date[2] := 19, [57].runs[0] := 6, [57].runs[17] := 1, [57].runs[18] := 2, [57].time_avg[0] := 112, [57].time_avg[2] := 41643, [57].time_avg[4] := 46281, [57].time_avg[5] := 22361, [57].time_avg[18] := 87, [58].date[0] := -2, [58].date[1] := 1, [58].date[2] := 15, [58].runs[0] := 7, [58].time_avg[0] := 126, [58].time_avg[4] := 37560, [58].time_avg[5] := 22361, [59].date[0] := -2, [59].date[1] := 1, [59].date[2] := 13, [59].runs[0] := 32, [59].runs[20] := 8, [59].runs[21] := 5, [59].runs[23] := 6, [59].time_avg[0] := 213,
        [59].time_avg[4] := 37560, [59].time_avg[5] := 22361, [59].time_avg[20] := 70, [59].time_avg[21] := 68, [59].time_avg[23] := 68, [60].date[0] := -2, [60].date[1] := 1, [60].date[2] := 12, [60].runs[0] := 17, [60].runs[20] := 5, [60].runs[21] := 5, [60].time_avg[0] := 121, [60].time_avg[4] := 37560, [60].time_avg[5] := 22361, [60].time_avg[20] := 167, [60].time_avg[21] := 64, [61].date[0] := -2, [61].date[1] := 1, [61].date[2] := 11, [61].runs[0] := 8, [61].runs[18] := 1, [61].runs[19] := 2, [61].runs[20] := 2, [61].runs[23] := 3, [61].time_avg[0] := 204, [61].time_avg[4] := 37560, [61].time_avg[5] := 22361, [61].time_avg[19] := 278, [61].time_avg[23] := 58, [62].date[0] := -2, [62].date[1] := 1, [62].date[2] := 10, [62].runs[0] := 4, [62].runs[18] := 1, [62].runs[20] := 2, [62].runs[23] := 1, [62].time_avg[0] := 4, [62].time_avg[2] := 30360, [62].time_avg[4] := 37560, [62].time_avg[5] := 22361, [62].time_avg[20] := 317, [63].date[0] := -2, [63].date[1] := 1, [63].date[2] := 8, [63].runs[0] := 28, [63].runs[17] := 1, [63].runs[18] := 1, [63].runs[20] := 4, [63].runs[21] := 2, [63].runs[23] := 3, [63].time_avg[0] := 184, [63].time_avg[2] := -4678, [63].time_avg[4] := 9800, [63].time_avg[5] := 22361, [63].time_avg[18] := 298, [63].time_avg[20] := 114, [63].time_avg[23] := 244, [64].date[0] := -2, [64].date[1] := 1, [64].date[2] := 7,
        [64].runs[0] := 9, [64].runs[17] := 1, [64].runs[19] := 1, [64].runs[20] := 3, [64].time_avg[0] := 370, [64].time_avg[5] := 22361, [64].time_avg[20] := 370, [65].date[0] := -2, [65].date[1] := 2, [65].date[2] := 10, [65].runs[0] := 14, [65].runs[19] := 9, [65].runs[20] := 5, [65].time_avg[5] := 22361, [66].date[0] := 20, [66].date[1] := 3, [66].date[2] := 5, [66].runs[0] := 11, [66].runs[8] := 1, [66].runs[9] := 1, [66].runs[10] := 1, [66].runs[14] := 3, [66].runs[15] := 1, [66].runs[16] := 2, [66].runs[17] := 2, [66].time_avg[0] := 250, [66].time_avg[5] := 22361, [66].time_avg[10] := 454, [66].time_avg[14] := 139, [66].time_avg[16] := 157, [67].date[0] := 20, [67].date[1] := 3, [67].date[2] := 4, [67].runs[0] := 20, [67].runs[11] := 4, [67].runs[12] := 6, [67].runs[18] := 8, [67].runs[19] := 2, [67].time_avg[0] := 36, [67].time_avg[2] := 31218, [67].time_avg[5] := 22361, [67].time_avg[12] := 36, [68].date[0] := 20, [68].date[1] := 3, [68].date[2] := 2, [68].runs[0] := 87, [68].runs[12] := 1, [68].runs[13] := 6, [68].runs[14] := 17, [68].runs[15] := 16, [68].runs[16] := 15, [68].runs[17] := 15, [68].runs[18] := 11, [68].runs[19] := 6, [68].time_avg[0] := 29, [68].time_avg[4] := 28480, [68].time_avg[5] := 22361, [68].time_avg[14] := 29, [68].time_avg[15] := 23, [68].time_avg[16] := 34,
